(* Logix 5000 project; controller FV vendor 1 type 14 code 217 rev 31.11; software revision 31.00; part 49 of 63 *)
(* tags used below, declared in another part *)
   CheckTimeMask : INT;
   CWD : CHECKWORD_FLAGS;
   Delphi_Does_Eng_Func : BOOL;
   FV_AV1 : PlantItem;   // AV1
   FV_AV1A : PlantItem;   // AV1A
   FV_AV2 : PlantItem;   // AV2
   FV_AV3 : PlantItem;   // AV3
   FV_AV4 : PlantItem;   // AV4
   FV_AV4A : PlantItem;   // AV4A
   FV_FV1C : PlantItem;   // FV1C
   FV_FV1J : PlantItem;   // FV1J
   FV_FV29C : PlantItem;   // FV29C
   FV_FV2C : PlantItem;   // FV2C
   FV_FV2J : PlantItem;   // FV2J
   FV_FV30C : PlantItem;   // FV30C
   FV_FV30J : PlantItem;   // FV30J
   FV_FV31C : PlantItem;   // FV31C
   FV_FV31J : PlantItem;   // FV31J
   FV_FV3C : PlantItem;   // FV3C
   FV_FV3J : PlantItem;   // FV3J
   FV_FV4C : PlantItem;   // FV4C
   FV_FV4J : PlantItem;   // FV4J
   FV_FV5C : PlantItem;   // FV5C
   FV_FV5J : PlantItem;   // FV5J
   FV_FV6C : PlantItem;   // FV6C
   FV_FV6J : PlantItem;   // FV6J
   FV_FV7C : PlantItem;   // FV7C
   FV_FV7J : PlantItem;   // FV7J
   FV_FV8C : PlantItem;   // FV8C
   FV_FV8J : PlantItem;   // FV8J
   FV_FV9C : PlantItem;   // FV9C
   FV_FV9J : PlantItem;   // FV9J
   FV_N255 : INT[255];   // Old Checkwords to keep Delphi working in the interim before full changeover.
   FV_R2V1 : PlantItem;   // R2V1
   FV_R2V2 : PlantItem;   // R2V2
   FV_WYT1R : PlantItem;   // WYT1R
   FV_WYT2R : PlantItem;   // WYT2R
   FV_WYTR1 : PlantItem;   // WYTR1
   FV_WYTR2 : PlantItem;   // WYTR2
   FV_YSV1R : PlantItem;   // YSV1R
   TempChecktime : DINT;
(* FV_Common, continued *)

   72: [XIC(Delphi_Does_Eng_Func) [[XIC(FV_N255[88].8) [OTL(FV_FV29C.CW.[CWD.MANUAL]) ,XIC(FV_N255[88].9) OTL(FV_FV29C.CW.[CWD.MANDRV]) ,XIO(FV_N255[88].9) OTU(FV_FV29C.CW.[CWD.MANDRV]) ] ,XIO(FV_N255[88].8) [OTU(FV_FV29C.CW.[CWD.MANUAL]) ,[XIC(FV_FV29C.CW.[CWD.OUTPUT]) OTL(FV_N255[88].9) ,XIO(FV_FV29C.CW.[CWD.OUTPUT]) OTU(FV_N255[88].9) ] ] ] ,[XIC(FV_N255[88].13) OTL(FV_FV29C.CW.[CWD.CHECKOFF]) ,XIO(FV_N255[88].13) OTU(FV_FV29C.CW.[CWD.CHECKOFF]) ] ] ,XIO(Delphi_Does_Eng_Func) [[XIC(FV_FV29C.CW.[CWD.MANUAL]) OTL(FV_N255[88].8) ,XIO(FV_FV29C.CW.[CWD.MANUAL]) OTU(FV_N255[88].8) ] ,[XIC(FV_FV29C.CW.[CWD.CHECKOFF]) OTL(FV_N255[88].13) ,XIO(FV_FV29C.CW.[CWD.CHECKOFF]) OTU(FV_N255[88].13) ] ,[XIC(FV_FV29C.CW.[CWD.OUTPUT]) OTL(FV_N255[88].9) ,XIO(FV_FV29C.CW.[CWD.OUTPUT]) OTU(FV_N255[88].9) ] ] ,XIC(FV_FV29C.CW.[CWD.OUTPUT]) OTE(FV_N255[88].10) ,XIO(FV_FV29C.CW.[CWD.OUTPUT]) OTE(FV_N255[88].11) ,XIC(FV_FV29C.CW.[CWD.FAULT]) OTE(FV_N255[88].15) ];
   73: [XIC(Delphi_Does_Eng_Func) [[XIC(FV_N255[89].8) [OTL(FV_FV30J.CW.[CWD.MANUAL]) ,XIC(FV_N255[89].9) OTL(FV_FV30J.CW.[CWD.MANDRV]) ,XIO(FV_N255[89].9) OTU(FV_FV30J.CW.[CWD.MANDRV]) ] ,XIO(FV_N255[89].8) [OTU(FV_FV30J.CW.[CWD.MANUAL]) ,[XIC(FV_FV30J.CW.[CWD.OUTPUT]) OTL(FV_N255[89].9) ,XIO(FV_FV30J.CW.[CWD.OUTPUT]) OTU(FV_N255[89].9) ] ] ] ,[XIC(FV_N255[89].13) OTL(FV_FV30J.CW.[CWD.CHECKOFF]) ,XIO(FV_N255[89].13) OTU(FV_FV30J.CW.[CWD.CHECKOFF]) ] ] ,XIO(Delphi_Does_Eng_Func) [[XIC(FV_FV30J.CW.[CWD.MANUAL]) OTL(FV_N255[89].8) ,XIO(FV_FV30J.CW.[CWD.MANUAL]) OTU(FV_N255[89].8) ] ,[XIC(FV_FV30J.CW.[CWD.CHECKOFF]) OTL(FV_N255[89].13) ,XIO(FV_FV30J.CW.[CWD.CHECKOFF]) OTU(FV_N255[89].13) ] ,[XIC(FV_FV30J.CW.[CWD.OUTPUT]) OTL(FV_N255[89].9) ,XIO(FV_FV30J.CW.[CWD.OUTPUT]) OTU(FV_N255[89].9) ] ] ,XIC(FV_FV30J.CW.[CWD.OUTPUT]) OTE(FV_N255[89].10) ,XIO(FV_FV30J.CW.[CWD.OUTPUT]) OTE(FV_N255[89].11) ,XIC(FV_FV30J.CW.[CWD.FAULT]) OTE(FV_N255[89].15) ];
   74: [XIC(Delphi_Does_Eng_Func) [[XIC(FV_N255[90].8) [OTL(FV_FV30C.CW.[CWD.MANUAL]) ,XIC(FV_N255[90].9) OTL(FV_FV30C.CW.[CWD.MANDRV]) ,XIO(FV_N255[90].9) OTU(FV_FV30C.CW.[CWD.MANDRV]) ] ,XIO(FV_N255[90].8) [OTU(FV_FV30C.CW.[CWD.MANUAL]) ,[XIC(FV_FV30C.CW.[CWD.OUTPUT]) OTL(FV_N255[90].9) ,XIO(FV_FV30C.CW.[CWD.OUTPUT]) OTU(FV_N255[90].9) ] ] ] ,[XIC(FV_N255[90].13) OTL(FV_FV30C.CW.[CWD.CHECKOFF]) ,XIO(FV_N255[90].13) OTU(FV_FV30C.CW.[CWD.CHECKOFF]) ] ] ,XIO(Delphi_Does_Eng_Func) [[XIC(FV_FV30C.CW.[CWD.MANUAL]) OTL(FV_N255[90].8) ,XIO(FV_FV30C.CW.[CWD.MANUAL]) OTU(FV_N255[90].8) ] ,[XIC(FV_FV30C.CW.[CWD.CHECKOFF]) OTL(FV_N255[90].13) ,XIO(FV_FV30C.CW.[CWD.CHECKOFF]) OTU(FV_N255[90].13) ] ,[XIC(FV_FV30C.CW.[CWD.OUTPUT]) OTL(FV_N255[90].9) ,XIO(FV_FV30C.CW.[CWD.OUTPUT]) OTU(FV_N255[90].9) ] ] ,XIC(FV_FV30C.CW.[CWD.OUTPUT]) OTE(FV_N255[90].10) ,XIO(FV_FV30C.CW.[CWD.OUTPUT]) OTE(FV_N255[90].11) ,XIC(FV_FV30C.CW.[CWD.FAULT]) OTE(FV_N255[90].15) ];
   75: [XIC(Delphi_Does_Eng_Func) [[XIC(FV_N255[91].8) [OTL(FV_FV31J.CW.[CWD.MANUAL]) ,XIC(FV_N255[91].9) OTL(FV_FV31J.CW.[CWD.MANDRV]) ,XIO(FV_N255[91].9) OTU(FV_FV31J.CW.[CWD.MANDRV]) ] ,XIO(FV_N255[91].8) [OTU(FV_FV31J.CW.[CWD.MANUAL]) ,[XIC(FV_FV31J.CW.[CWD.OUTPUT]) OTL(FV_N255[91].9) ,XIO(FV_FV31J.CW.[CWD.OUTPUT]) OTU(FV_N255[91].9) ] ] ] ,[XIC(FV_N255[91].13) OTL(FV_FV31J.CW.[CWD.CHECKOFF]) ,XIO(FV_N255[91].13) OTU(FV_FV31J.CW.[CWD.CHECKOFF]) ] ] ,XIO(Delphi_Does_Eng_Func) [[XIC(FV_FV31J.CW.[CWD.MANUAL]) OTL(FV_N255[91].8) ,XIO(FV_FV31J.CW.[CWD.MANUAL]) OTU(FV_N255[91].8) ] ,[XIC(FV_FV31J.CW.[CWD.CHECKOFF]) OTL(FV_N255[91].13) ,XIO(FV_FV31J.CW.[CWD.CHECKOFF]) OTU(FV_N255[91].13) ] ,[XIC(FV_FV31J.CW.[CWD.OUTPUT]) OTL(FV_N255[91].9) ,XIO(FV_FV31J.CW.[CWD.OUTPUT]) OTU(FV_N255[91].9) ] ] ,XIC(FV_FV31J.CW.[CWD.OUTPUT]) OTE(FV_N255[91].10) ,XIO(FV_FV31J.CW.[CWD.OUTPUT]) OTE(FV_N255[91].11) ,XIC(FV_FV31J.CW.[CWD.FAULT]) OTE(FV_N255[91].15) ];
   76: [XIC(Delphi_Does_Eng_Func) [[XIC(FV_N255[92].8) [OTL(FV_FV31C.CW.[CWD.MANUAL]) ,XIC(FV_N255[92].9) OTL(FV_FV31C.CW.[CWD.MANDRV]) ,XIO(FV_N255[92].9) OTU(FV_FV31C.CW.[CWD.MANDRV]) ] ,XIO(FV_N255[92].8) [OTU(FV_FV31C.CW.[CWD.MANUAL]) ,[XIC(FV_FV31C.CW.[CWD.OUTPUT]) OTL(FV_N255[92].9) ,XIO(FV_FV31C.CW.[CWD.OUTPUT]) OTU(FV_N255[92].9) ] ] ] ,[XIC(FV_N255[92].13) OTL(FV_FV31C.CW.[CWD.CHECKOFF]) ,XIO(FV_N255[92].13) OTU(FV_FV31C.CW.[CWD.CHECKOFF]) ] ] ,XIO(Delphi_Does_Eng_Func) [[XIC(FV_FV31C.CW.[CWD.MANUAL]) OTL(FV_N255[92].8) ,XIO(FV_FV31C.CW.[CWD.MANUAL]) OTU(FV_N255[92].8) ] ,[XIC(FV_FV31C.CW.[CWD.CHECKOFF]) OTL(FV_N255[92].13) ,XIO(FV_FV31C.CW.[CWD.CHECKOFF]) OTU(FV_N255[92].13) ] ,[XIC(FV_FV31C.CW.[CWD.OUTPUT]) OTL(FV_N255[92].9) ,XIO(FV_FV31C.CW.[CWD.OUTPUT]) OTU(FV_N255[92].9) ] ] ,XIC(FV_FV31C.CW.[CWD.OUTPUT]) OTE(FV_N255[92].10) ,XIO(FV_FV31C.CW.[CWD.OUTPUT]) OTE(FV_N255[92].11) ,XIC(FV_FV31C.CW.[CWD.FAULT]) OTE(FV_N255[92].15) ];
   77: [XIC(Delphi_Does_Eng_Func) [[XIC(FV_N255[79].8) [OTL(FV_WYT1R.CW.[CWD.MANUAL]) ,XIC(FV_N255[79].9) OTL(FV_WYT1R.CW.[CWD.MANDRV]) ,XIO(FV_N255[79].9) OTU(FV_WYT1R.CW.[CWD.MANDRV]) ] ,XIO(FV_N255[79].8) [OTU(FV_WYT1R.CW.[CWD.MANUAL]) ,[XIC(FV_WYT1R.CW.[CWD.OUTPUT]) OTL(FV_N255[79].9) ,XIO(FV_WYT1R.CW.[CWD.OUTPUT]) OTU(FV_N255[79].9) ] ] ] ,[XIC(FV_N255[79].13) OTL(FV_WYT1R.CW.[CWD.CHECKOFF]) ,XIO(FV_N255[79].13) OTU(FV_WYT1R.CW.[CWD.CHECKOFF]) ] ] ,XIO(Delphi_Does_Eng_Func) [[XIC(FV_WYT1R.CW.[CWD.MANUAL]) OTL(FV_N255[79].8) ,XIO(FV_WYT1R.CW.[CWD.MANUAL]) OTU(FV_N255[79].8) ] ,[XIC(FV_WYT1R.CW.[CWD.CHECKOFF]) OTL(FV_N255[79].13) ,XIO(FV_WYT1R.CW.[CWD.CHECKOFF]) OTU(FV_N255[79].13) ] ,[XIC(FV_WYT1R.CW.[CWD.OUTPUT]) OTL(FV_N255[79].9) ,XIO(FV_WYT1R.CW.[CWD.OUTPUT]) OTU(FV_N255[79].9) ] ] ,XIC(FV_WYT1R.CW.[CWD.RUNFB]) OTE(FV_N255[79].10) ,XIO(FV_WYT1R.CW.[CWD.RUNFB]) OTE(FV_N255[79].11) ,XIC(FV_WYT1R.CW.[CWD.FAULT]) OTE(FV_N255[79].15) ];
   78: [XIC(Delphi_Does_Eng_Func) [[XIC(FV_N255[80].8) [OTL(FV_WYT2R.CW.[CWD.MANUAL]) ,XIC(FV_N255[80].9) OTL(FV_WYT2R.CW.[CWD.MANDRV]) ,XIO(FV_N255[80].9) OTU(FV_WYT2R.CW.[CWD.MANDRV]) ] ,XIO(FV_N255[80].8) [OTU(FV_WYT2R.CW.[CWD.MANUAL]) ,[XIC(FV_WYT2R.CW.[CWD.OUTPUT]) OTL(FV_N255[80].9) ,XIO(FV_WYT2R.CW.[CWD.OUTPUT]) OTU(FV_N255[80].9) ] ] ] ,[XIC(FV_N255[80].13) OTL(FV_WYT2R.CW.[CWD.CHECKOFF]) ,XIO(FV_N255[80].13) OTU(FV_WYT2R.CW.[CWD.CHECKOFF]) ] ] ,XIO(Delphi_Does_Eng_Func) [[XIC(FV_WYT2R.CW.[CWD.MANUAL]) OTL(FV_N255[80].8) ,XIO(FV_WYT2R.CW.[CWD.MANUAL]) OTU(FV_N255[80].8) ] ,[XIC(FV_WYT2R.CW.[CWD.CHECKOFF]) OTL(FV_N255[80].13) ,XIO(FV_WYT2R.CW.[CWD.CHECKOFF]) OTU(FV_N255[80].13) ] ,[XIC(FV_WYT2R.CW.[CWD.OUTPUT]) OTL(FV_N255[80].9) ,XIO(FV_WYT2R.CW.[CWD.OUTPUT]) OTU(FV_N255[80].9) ] ] ,XIC(FV_WYT2R.CW.[CWD.RUNFB]) OTE(FV_N255[80].10) ,XIO(FV_WYT2R.CW.[CWD.RUNFB]) OTE(FV_N255[80].11) ,XIC(FV_WYT2R.CW.[CWD.FAULT]) OTE(FV_N255[80].15) ];
   79: [XIC(Delphi_Does_Eng_Func) [[XIC(FV_N255[59].8) [OTL(FV_YSV1R.CW.[CWD.MANUAL]) ,XIC(FV_N255[59].9) OTL(FV_YSV1R.CW.[CWD.MANDRV]) ,XIO(FV_N255[59].9) OTU(FV_YSV1R.CW.[CWD.MANDRV]) ] ,XIO(FV_N255[59].8) [OTU(FV_YSV1R.CW.[CWD.MANUAL]) ,[XIC(FV_YSV1R.CW.[CWD.OUTPUT]) OTL(FV_N255[59].9) ,XIO(FV_YSV1R.CW.[CWD.OUTPUT]) OTU(FV_N255[59].9) ] ] ] ,[XIC(FV_N255[59].13) OTL(FV_YSV1R.CW.[CWD.CHECKOFF]) ,XIO(FV_N255[59].13) OTU(FV_YSV1R.CW.[CWD.CHECKOFF]) ] ] ,XIO(Delphi_Does_Eng_Func) [[XIC(FV_YSV1R.CW.[CWD.MANUAL]) OTL(FV_N255[59].8) ,XIO(FV_YSV1R.CW.[CWD.MANUAL]) OTU(FV_N255[59].8) ] ,[XIC(FV_YSV1R.CW.[CWD.CHECKOFF]) OTL(FV_N255[59].13) ,XIO(FV_YSV1R.CW.[CWD.CHECKOFF]) OTU(FV_N255[59].13) ] ,[XIC(FV_YSV1R.CW.[CWD.OUTPUT]) OTL(FV_N255[59].9) ,XIO(FV_YSV1R.CW.[CWD.OUTPUT]) OTU(FV_N255[59].9) ] ] ,XIC(FV_YSV1R.CW.[CWD.RUNFB]) OTE(FV_N255[59].10) ,XIO(FV_YSV1R.CW.[CWD.RUNFB]) OTE(FV_N255[59].11) ,XIC(FV_YSV1R.CW.[CWD.FAULT]) OTE(FV_N255[59].15) ];
   80: [XIC(Delphi_Does_Eng_Func) [[XIC(FV_N255[65].8) [OTL(FV_AV1.CW.[CWD.MANUAL]) ,XIC(FV_N255[65].9) OTL(FV_AV1.CW.[CWD.MANDRV]) ,XIO(FV_N255[65].9) OTU(FV_AV1.CW.[CWD.MANDRV]) ] ,XIO(FV_N255[65].8) [OTU(FV_AV1.CW.[CWD.MANUAL]) ,[XIC(FV_AV1.CW.[CWD.OUTPUT]) OTL(FV_N255[65].9) ,XIO(FV_AV1.CW.[CWD.OUTPUT]) OTU(FV_N255[65].9) ] ] ] ,[XIC(FV_N255[65].13) OTL(FV_AV1.CW.[CWD.CHECKOFF]) ,XIO(FV_N255[65].13) OTU(FV_AV1.CW.[CWD.CHECKOFF]) ] ] ,XIO(Delphi_Does_Eng_Func) [[XIC(FV_AV1.CW.[CWD.MANUAL]) OTL(FV_N255[65].8) ,XIO(FV_AV1.CW.[CWD.MANUAL]) OTU(FV_N255[65].8) ] ,[XIC(FV_AV1.CW.[CWD.CHECKOFF]) OTL(FV_N255[65].13) ,XIO(FV_AV1.CW.[CWD.CHECKOFF]) OTU(FV_N255[65].13) ] ,[XIC(FV_AV1.CW.[CWD.OUTPUT]) OTL(FV_N255[65].9) ,XIO(FV_AV1.CW.[CWD.OUTPUT]) OTU(FV_N255[65].9) ] ] ,XIC(FV_AV1.CW.[CWD.OPENFB]) OTE(FV_N255[65].10) ,XIC(FV_AV1.CW.[CWD.CLOSEDFB]) OTE(FV_N255[65].11) ,XIC(FV_AV1.CW.[CWD.FAULT]) OTE(FV_N255[65].15) ];
   81: [XIC(Delphi_Does_Eng_Func) [[XIC(FV_N255[66].8) [OTL(FV_AV2.CW.[CWD.MANUAL]) ,XIC(FV_N255[66].9) OTL(FV_AV2.CW.[CWD.MANDRV]) ,XIO(FV_N255[66].9) OTU(FV_AV2.CW.[CWD.MANDRV]) ] ,XIO(FV_N255[66].8) [OTU(FV_AV2.CW.[CWD.MANUAL]) ,[XIC(FV_AV2.CW.[CWD.OUTPUT]) OTL(FV_N255[66].9) ,XIO(FV_AV2.CW.[CWD.OUTPUT]) OTU(FV_N255[66].9) ] ] ] ,[XIC(FV_N255[66].13) OTL(FV_AV2.CW.[CWD.CHECKOFF]) ,XIO(FV_N255[66].13) OTU(FV_AV2.CW.[CWD.CHECKOFF]) ] ] ,XIO(Delphi_Does_Eng_Func) [[XIC(FV_AV2.CW.[CWD.MANUAL]) OTL(FV_N255[66].8) ,XIO(FV_AV2.CW.[CWD.MANUAL]) OTU(FV_N255[66].8) ] ,[XIC(FV_AV2.CW.[CWD.CHECKOFF]) OTL(FV_N255[66].13) ,XIO(FV_AV2.CW.[CWD.CHECKOFF]) OTU(FV_N255[66].13) ] ,[XIC(FV_AV2.CW.[CWD.OUTPUT]) OTL(FV_N255[66].9) ,XIO(FV_AV2.CW.[CWD.OUTPUT]) OTU(FV_N255[66].9) ] ] ,XIC(FV_AV2.CW.[CWD.OPENFB]) OTE(FV_N255[66].10) ,XIC(FV_AV2.CW.[CWD.CLOSEDFB]) OTE(FV_N255[66].11) ,XIC(FV_AV2.CW.[CWD.FAULT]) OTE(FV_N255[66].15) ];
   82: [XIC(Delphi_Does_Eng_Func) [[XIC(FV_N255[67].8) [OTL(FV_AV3.CW.[CWD.MANUAL]) ,XIC(FV_N255[67].9) OTL(FV_AV3.CW.[CWD.MANDRV]) ,XIO(FV_N255[67].9) OTU(FV_AV3.CW.[CWD.MANDRV]) ] ,XIO(FV_N255[67].8) [OTU(FV_AV3.CW.[CWD.MANUAL]) ,[XIC(FV_AV3.CW.[CWD.OUTPUT]) OTL(FV_N255[67].9) ,XIO(FV_AV3.CW.[CWD.OUTPUT]) OTU(FV_N255[67].9) ] ] ] ,[XIC(FV_N255[67].13) OTL(FV_AV3.CW.[CWD.CHECKOFF]) ,XIO(FV_N255[67].13) OTU(FV_AV3.CW.[CWD.CHECKOFF]) ] ] ,XIO(Delphi_Does_Eng_Func) [[XIC(FV_AV3.CW.[CWD.MANUAL]) OTL(FV_N255[67].8) ,XIO(FV_AV3.CW.[CWD.MANUAL]) OTU(FV_N255[67].8) ] ,[XIC(FV_AV3.CW.[CWD.CHECKOFF]) OTL(FV_N255[67].13) ,XIO(FV_AV3.CW.[CWD.CHECKOFF]) OTU(FV_N255[67].13) ] ,[XIC(FV_AV3.CW.[CWD.OUTPUT]) OTL(FV_N255[67].9) ,XIO(FV_AV3.CW.[CWD.OUTPUT]) OTU(FV_N255[67].9) ] ] ,XIC(FV_AV3.CW.[CWD.OPENFB]) OTE(FV_N255[67].10) ,XIC(FV_AV3.CW.[CWD.CLOSEDFB]) OTE(FV_N255[67].11) ,XIC(FV_AV3.CW.[CWD.FAULT]) OTE(FV_N255[67].15) ];
   83: [XIC(Delphi_Does_Eng_Func) [[XIC(FV_N255[68].8) [OTL(FV_AV4.CW.[CWD.MANUAL]) ,XIC(FV_N255[68].9) OTL(FV_AV4.CW.[CWD.MANDRV]) ,XIO(FV_N255[68].9) OTU(FV_AV4.CW.[CWD.MANDRV]) ] ,XIO(FV_N255[68].8) [OTU(FV_AV4.CW.[CWD.MANUAL]) ,[XIC(FV_AV4.CW.[CWD.OUTPUT]) OTL(FV_N255[68].9) ,XIO(FV_AV4.CW.[CWD.OUTPUT]) OTU(FV_N255[68].9) ] ] ] ,[XIC(FV_N255[68].13) OTL(FV_AV4.CW.[CWD.CHECKOFF]) ,XIO(FV_N255[68].13) OTU(FV_AV4.CW.[CWD.CHECKOFF]) ] ] ,XIO(Delphi_Does_Eng_Func) [[XIC(FV_AV4.CW.[CWD.MANUAL]) OTL(FV_N255[68].8) ,XIO(FV_AV4.CW.[CWD.MANUAL]) OTU(FV_N255[68].8) ] ,[XIC(FV_AV4.CW.[CWD.CHECKOFF]) OTL(FV_N255[68].13) ,XIO(FV_AV4.CW.[CWD.CHECKOFF]) OTU(FV_N255[68].13) ] ,[XIC(FV_AV4.CW.[CWD.OUTPUT]) OTL(FV_N255[68].9) ,XIO(FV_AV4.CW.[CWD.OUTPUT]) OTU(FV_N255[68].9) ] ] ,XIC(FV_AV4.CW.[CWD.OPENFB]) OTE(FV_N255[68].10) ,XIC(FV_AV4.CW.[CWD.CLOSEDFB]) OTE(FV_N255[68].11) ,XIC(FV_AV4.CW.[CWD.FAULT]) OTE(FV_N255[68].15) ];
   84: [XIC(Delphi_Does_Eng_Func) [[XIC(FV_N255[69].8) [OTL(FV_AV1A.CW.[CWD.MANUAL]) ,XIC(FV_N255[69].9) OTL(FV_AV1A.CW.[CWD.MANDRV]) ,XIO(FV_N255[69].9) OTU(FV_AV1A.CW.[CWD.MANDRV]) ] ,XIO(FV_N255[69].8) [OTU(FV_AV1A.CW.[CWD.MANUAL]) ,[XIC(FV_AV1A.CW.[CWD.OUTPUT]) OTL(FV_N255[69].9) ,XIO(FV_AV1A.CW.[CWD.OUTPUT]) OTU(FV_N255[69].9) ] ] ] ,[XIC(FV_N255[69].13) OTL(FV_AV1A.CW.[CWD.CHECKOFF]) ,XIO(FV_N255[69].13) OTU(FV_AV1A.CW.[CWD.CHECKOFF]) ] ] ,XIO(Delphi_Does_Eng_Func) [[XIC(FV_AV1A.CW.[CWD.MANUAL]) OTL(FV_N255[69].8) ,XIO(FV_AV1A.CW.[CWD.MANUAL]) OTU(FV_N255[69].8) ] ,[XIC(FV_AV1A.CW.[CWD.CHECKOFF]) OTL(FV_N255[69].13) ,XIO(FV_AV1A.CW.[CWD.CHECKOFF]) OTU(FV_N255[69].13) ] ,[XIC(FV_AV1A.CW.[CWD.OUTPUT]) OTL(FV_N255[69].9) ,XIO(FV_AV1A.CW.[CWD.OUTPUT]) OTU(FV_N255[69].9) ] ] ,XIC(FV_AV1A.CW.[CWD.OPENFB]) OTE(FV_N255[69].10) ,XIC(FV_AV1A.CW.[CWD.CLOSEDFB]) OTE(FV_N255[69].11) ,XIC(FV_AV1A.CW.[CWD.FAULT]) OTE(FV_N255[69].15) ];
   85: [XIC(Delphi_Does_Eng_Func) [[XIC(FV_N255[70].8) [OTL(FV_AV4A.CW.[CWD.MANUAL]) ,XIC(FV_N255[70].9) OTL(FV_AV4A.CW.[CWD.MANDRV]) ,XIO(FV_N255[70].9) OTU(FV_AV4A.CW.[CWD.MANDRV]) ] ,XIO(FV_N255[70].8) [OTU(FV_AV4A.CW.[CWD.MANUAL]) ,[XIC(FV_AV4A.CW.[CWD.OUTPUT]) OTL(FV_N255[70].9) ,XIO(FV_AV4A.CW.[CWD.OUTPUT]) OTU(FV_N255[70].9) ] ] ] ,[XIC(FV_N255[70].13) OTL(FV_AV4A.CW.[CWD.CHECKOFF]) ,XIO(FV_N255[70].13) OTU(FV_AV4A.CW.[CWD.CHECKOFF]) ] ] ,XIO(Delphi_Does_Eng_Func) [[XIC(FV_AV4A.CW.[CWD.MANUAL]) OTL(FV_N255[70].8) ,XIO(FV_AV4A.CW.[CWD.MANUAL]) OTU(FV_N255[70].8) ] ,[XIC(FV_AV4A.CW.[CWD.CHECKOFF]) OTL(FV_N255[70].13) ,XIO(FV_AV4A.CW.[CWD.CHECKOFF]) OTU(FV_N255[70].13) ] ,[XIC(FV_AV4A.CW.[CWD.OUTPUT]) OTL(FV_N255[70].9) ,XIO(FV_AV4A.CW.[CWD.OUTPUT]) OTU(FV_N255[70].9) ] ] ,XIC(FV_AV4A.CW.[CWD.OPENFB]) OTE(FV_N255[70].10) ,XIC(FV_AV4A.CW.[CWD.CLOSEDFB]) OTE(FV_N255[70].11) ,XIC(FV_AV4A.CW.[CWD.FAULT]) OTE(FV_N255[70].15) ];
   86: [XIC(Delphi_Does_Eng_Func) [[XIC(FV_N255[73].8) [OTL(FV_WYTR1.CW.[CWD.MANUAL]) ,XIC(FV_N255[73].9) OTL(FV_WYTR1.CW.[CWD.MANDRV]) ,XIO(FV_N255[73].9) OTU(FV_WYTR1.CW.[CWD.MANDRV]) ] ,XIO(FV_N255[73].8) [OTU(FV_WYTR1.CW.[CWD.MANUAL]) ,[XIC(FV_WYTR1.CW.[CWD.OUTPUT]) OTL(FV_N255[73].9) ,XIO(FV_WYTR1.CW.[CWD.OUTPUT]) OTU(FV_N255[73].9) ] ] ] ,[XIC(FV_N255[73].13) OTL(FV_WYTR1.CW.[CWD.CHECKOFF]) ,XIO(FV_N255[73].13) OTU(FV_WYTR1.CW.[CWD.CHECKOFF]) ] ] ,XIO(Delphi_Does_Eng_Func) [[XIC(FV_WYTR1.CW.[CWD.MANUAL]) OTL(FV_N255[73].8) ,XIO(FV_WYTR1.CW.[CWD.MANUAL]) OTU(FV_N255[73].8) ] ,[XIC(FV_WYTR1.CW.[CWD.CHECKOFF]) OTL(FV_N255[73].13) ,XIO(FV_WYTR1.CW.[CWD.CHECKOFF]) OTU(FV_N255[73].13) ] ,[XIC(FV_WYTR1.CW.[CWD.OUTPUT]) OTL(FV_N255[73].9) ,XIO(FV_WYTR1.CW.[CWD.OUTPUT]) OTU(FV_N255[73].9) ] ] ,XIC(FV_WYTR1.CW.[CWD.OPENFB]) OTE(FV_N255[73].10) ,XIC(FV_WYTR1.CW.[CWD.CLOSEDFB]) OTE(FV_N255[73].11) ,XIC(FV_WYTR1.CW.[CWD.FAULT]) OTE(FV_N255[73].15) ];
   87: [XIC(Delphi_Does_Eng_Func) [[XIC(FV_N255[74].8) [OTL(FV_WYTR2.CW.[CWD.MANUAL]) ,XIC(FV_N255[74].9) OTL(FV_WYTR2.CW.[CWD.MANDRV]) ,XIO(FV_N255[74].9) OTU(FV_WYTR2.CW.[CWD.MANDRV]) ] ,XIO(FV_N255[74].8) [OTU(FV_WYTR2.CW.[CWD.MANUAL]) ,[XIC(FV_WYTR2.CW.[CWD.OUTPUT]) OTL(FV_N255[74].9) ,XIO(FV_WYTR2.CW.[CWD.OUTPUT]) OTU(FV_N255[74].9) ] ] ] ,[XIC(FV_N255[74].13) OTL(FV_WYTR2.CW.[CWD.CHECKOFF]) ,XIO(FV_N255[74].13) OTU(FV_WYTR2.CW.[CWD.CHECKOFF]) ] ] ,XIO(Delphi_Does_Eng_Func) [[XIC(FV_WYTR2.CW.[CWD.MANUAL]) OTL(FV_N255[74].8) ,XIO(FV_WYTR2.CW.[CWD.MANUAL]) OTU(FV_N255[74].8) ] ,[XIC(FV_WYTR2.CW.[CWD.CHECKOFF]) OTL(FV_N255[74].13) ,XIO(FV_WYTR2.CW.[CWD.CHECKOFF]) OTU(FV_N255[74].13) ] ,[XIC(FV_WYTR2.CW.[CWD.OUTPUT]) OTL(FV_N255[74].9) ,XIO(FV_WYTR2.CW.[CWD.OUTPUT]) OTU(FV_N255[74].9) ] ] ,XIC(FV_WYTR2.CW.[CWD.OPENFB]) OTE(FV_N255[74].10) ,XIC(FV_WYTR2.CW.[CWD.CLOSEDFB]) OTE(FV_N255[74].11) ,XIC(FV_WYTR2.CW.[CWD.FAULT]) OTE(FV_N255[74].15) ];
   88: [XIC(Delphi_Does_Eng_Func) [[XIC(FV_N255[75].8) [OTL(FV_R2V1.CW.[CWD.MANUAL]) ,XIC(FV_N255[75].9) OTL(FV_R2V1.CW.[CWD.MANDRV]) ,XIO(FV_N255[75].9) OTU(FV_R2V1.CW.[CWD.MANDRV]) ] ,XIO(FV_N255[75].8) [OTU(FV_R2V1.CW.[CWD.MANUAL]) ,[XIC(FV_R2V1.CW.[CWD.OUTPUT]) OTL(FV_N255[75].9) ,XIO(FV_R2V1.CW.[CWD.OUTPUT]) OTU(FV_N255[75].9) ] ] ] ,[XIC(FV_N255[75].13) OTL(FV_R2V1.CW.[CWD.CHECKOFF]) ,XIO(FV_N255[75].13) OTU(FV_R2V1.CW.[CWD.CHECKOFF]) ] ] ,XIO(Delphi_Does_Eng_Func) [[XIC(FV_R2V1.CW.[CWD.MANUAL]) OTL(FV_N255[75].8) ,XIO(FV_R2V1.CW.[CWD.MANUAL]) OTU(FV_N255[75].8) ] ,[XIC(FV_R2V1.CW.[CWD.CHECKOFF]) OTL(FV_N255[75].13) ,XIO(FV_R2V1.CW.[CWD.CHECKOFF]) OTU(FV_N255[75].13) ] ,[XIC(FV_R2V1.CW.[CWD.OUTPUT]) OTL(FV_N255[75].9) ,XIO(FV_R2V1.CW.[CWD.OUTPUT]) OTU(FV_N255[75].9) ] ] ,XIC(FV_R2V1.CW.[CWD.OPENFB]) OTE(FV_N255[75].10) ,XIC(FV_R2V1.CW.[CWD.CLOSEDFB]) OTE(FV_N255[75].11) ,XIC(FV_R2V1.CW.[CWD.FAULT]) OTE(FV_N255[75].15) ];
   89: [XIC(Delphi_Does_Eng_Func) [[XIC(FV_N255[76].8) [OTL(FV_R2V2.CW.[CWD.MANUAL]) ,XIC(FV_N255[76].9) OTL(FV_R2V2.CW.[CWD.MANDRV]) ,XIO(FV_N255[76].9) OTU(FV_R2V2.CW.[CWD.MANDRV]) ] ,XIO(FV_N255[76].8) [OTU(FV_R2V2.CW.[CWD.MANUAL]) ,[XIC(FV_R2V2.CW.[CWD.OUTPUT]) OTL(FV_N255[76].9) ,XIO(FV_R2V2.CW.[CWD.OUTPUT]) OTU(FV_N255[76].9) ] ] ] ,[XIC(FV_N255[76].13) OTL(FV_R2V2.CW.[CWD.CHECKOFF]) ,XIO(FV_N255[76].13) OTU(FV_R2V2.CW.[CWD.CHECKOFF]) ] ] ,XIO(Delphi_Does_Eng_Func) [[XIC(FV_R2V2.CW.[CWD.MANUAL]) OTL(FV_N255[76].8) ,XIO(FV_R2V2.CW.[CWD.MANUAL]) OTU(FV_N255[76].8) ] ,[XIC(FV_R2V2.CW.[CWD.CHECKOFF]) OTL(FV_N255[76].13) ,XIO(FV_R2V2.CW.[CWD.CHECKOFF]) OTU(FV_N255[76].13) ] ,[XIC(FV_R2V2.CW.[CWD.OUTPUT]) OTL(FV_N255[76].9) ,XIO(FV_R2V2.CW.[CWD.OUTPUT]) OTU(FV_N255[76].9) ] ] ,XIC(FV_R2V2.CW.[CWD.OPENFB]) OTE(FV_N255[76].10) ,XIC(FV_R2V2.CW.[CWD.CLOSEDFB]) OTE(FV_N255[76].11) ,XIC(FV_R2V2.CW.[CWD.FAULT]) OTE(FV_N255[76].15) ];
   90: XIC(Delphi_Does_Eng_Func)AND(FV_N255[1],CheckTimeMask,TempChecktime)[GRT(TempChecktime,0) DIV(TempChecktime,8,FV_FV1C.CheckTime) ,EQU(TempChecktime,0) OTL(FV_N255[1].6) ];
   91: XIC(Delphi_Does_Eng_Func)AND(FV_N255[2],CheckTimeMask,TempChecktime)[GRT(TempChecktime,0) DIV(TempChecktime,8,FV_FV1J.CheckTime) ,EQU(TempChecktime,0) OTL(FV_N255[2].6) ];
   92: XIC(Delphi_Does_Eng_Func)AND(FV_N255[3],CheckTimeMask,TempChecktime)[GRT(TempChecktime,0) DIV(TempChecktime,8,FV_FV2C.CheckTime) ,EQU(TempChecktime,0) OTL(FV_N255[3].6) ];
   93: XIC(Delphi_Does_Eng_Func)AND(FV_N255[4],CheckTimeMask,TempChecktime)[GRT(TempChecktime,0) DIV(TempChecktime,8,FV_FV2J.CheckTime) ,EQU(TempChecktime,0) OTL(FV_N255[4].6) ];
   94: XIC(Delphi_Does_Eng_Func)AND(FV_N255[5],CheckTimeMask,TempChecktime)[GRT(TempChecktime,0) DIV(TempChecktime,8,FV_FV3C.CheckTime) ,EQU(TempChecktime,0) OTL(FV_N255[5].6) ];
   95: XIC(Delphi_Does_Eng_Func)AND(FV_N255[6],CheckTimeMask,TempChecktime)[GRT(TempChecktime,0) DIV(TempChecktime,8,FV_FV3J.CheckTime) ,EQU(TempChecktime,0) OTL(FV_N255[6].6) ];
   96: XIC(Delphi_Does_Eng_Func)AND(FV_N255[7],CheckTimeMask,TempChecktime)[GRT(TempChecktime,0) DIV(TempChecktime,8,FV_FV4C.CheckTime) ,EQU(TempChecktime,0) OTL(FV_N255[7].6) ];
   97: XIC(Delphi_Does_Eng_Func)AND(FV_N255[8],CheckTimeMask,TempChecktime)[GRT(TempChecktime,0) DIV(TempChecktime,8,FV_FV4J.CheckTime) ,EQU(TempChecktime,0) OTL(FV_N255[8].6) ];
   98: XIC(Delphi_Does_Eng_Func)AND(FV_N255[9],CheckTimeMask,TempChecktime)[GRT(TempChecktime,0) DIV(TempChecktime,8,FV_FV5C.CheckTime) ,EQU(TempChecktime,0) OTL(FV_N255[9].6) ];
   99: XIC(Delphi_Does_Eng_Func)AND(FV_N255[10],CheckTimeMask,TempChecktime)[GRT(TempChecktime,0) DIV(TempChecktime,8,FV_FV5J.CheckTime) ,EQU(TempChecktime,0) OTL(FV_N255[10].6) ];
   100: XIC(Delphi_Does_Eng_Func)AND(FV_N255[11],CheckTimeMask,TempChecktime)[GRT(TempChecktime,0) DIV(TempChecktime,8,FV_FV6C.CheckTime) ,EQU(TempChecktime,0) OTL(FV_N255[11].6) ];
   101: XIC(Delphi_Does_Eng_Func)AND(FV_N255[12],CheckTimeMask,TempChecktime)[GRT(TempChecktime,0) DIV(TempChecktime,8,FV_FV6J.CheckTime) ,EQU(TempChecktime,0) OTL(FV_N255[12].6) ];
   102: XIC(Delphi_Does_Eng_Func)AND(FV_N255[13],CheckTimeMask,TempChecktime)[GRT(TempChecktime,0) DIV(TempChecktime,8,FV_FV7C.CheckTime) ,EQU(TempChecktime,0) OTL(FV_N255[13].6) ];
   103: XIC(Delphi_Does_Eng_Func)AND(FV_N255[14],CheckTimeMask,TempChecktime)[GRT(TempChecktime,0) DIV(TempChecktime,8,FV_FV7J.CheckTime) ,EQU(TempChecktime,0) OTL(FV_N255[14].6) ];
   104: XIC(Delphi_Does_Eng_Func)AND(FV_N255[15],CheckTimeMask,TempChecktime)[GRT(TempChecktime,0) DIV(TempChecktime,8,FV_FV8C.CheckTime) ,EQU(TempChecktime,0) OTL(FV_N255[15].6) ];
   105: XIC(Delphi_Does_Eng_Func)AND(FV_N255[16],CheckTimeMask,TempChecktime)[GRT(TempChecktime,0) DIV(TempChecktime,8,FV_FV8J.CheckTime) ,EQU(TempChecktime,0) OTL(FV_N255[16].6) ];
   106: XIC(Delphi_Does_Eng_Func)AND(FV_N255[17],CheckTimeMask,TempChecktime)[GRT(TempChecktime,0) DIV(TempChecktime,8,FV_FV9C.CheckTime) ,EQU(TempChecktime,0) OTL(FV_N255[17].6) ];
   107: XIC(Delphi_Does_Eng_Func)AND(FV_N255[18],CheckTimeMask,TempChecktime)[GRT(TempChecktime,0) DIV(TempChecktime,8,FV_FV9J.CheckTime) ,EQU(TempChecktime,0) OTL(FV_N255[18].6) ];
